// TIA Portal project "OPA_Demo" (V13)

(* hardware
DEVICE "S7-1200 station_1"  S7-1200 Station
   slot 0: "Rack_0"  Rack  V1.0
   slot 1: "PLC_1"  CPU 1214C DC/DC/DC  6ES7 214-1AG31-0XB0  V3.0
DEVICE "HMI_1"  KTP600 Basic color PN
   slot 0: "HMI"  HMI  6AV6 647-0AD11-3AX0  12.0.0.0
   slot 1: "HMI_RT_1"  KTP600 Basic color PN  6AV6 647-0AD11-3AX0  12.0.0.0
   slot 5: "HMI_1.IE_CP_1"  PROFINET Interface
      slot 1: "PROFINET Interface_1"  PROFINET Interface
         slot 1: "Port_1"  Port
*)

// ===== PLC "PLC_1"  CPU 1214C DC/DC/DC =====

VAR_GLOBAL   // PLC tag table "Input"
   "Tray_sensor" AT %I0.0 : Bool;
   "Doos_sensor" AT %I0.6 : Bool;
   "Tafel_sensor" AT %I0.4 : Bool;
   "Noodstop_aan_Plc" AT %I0.5 : Bool;
   "Noodstop_extern" AT %I0.3 : Bool;
   "Skip_Camera_Knop" AT %I0.1 : Bool;
   "Pause_Knop" AT %I0.2 : Bool;
END_VAR

VAR_GLOBAL   // PLC tag table "Memory"
   "HMI_Start_Pressed" AT %M42.0 : Bool;
   "HMI_Stop_Pressed" AT %M42.1 : Bool;
   "Running" AT %M42.2 : Bool;
   "HMI_White_Selected" AT %M42.3 : Bool;
   "HMI_Black_Pressed" AT %M42.4 : Bool;
   "HMI_tafel_omhoog" AT %M43.0 : Bool;
   "HMI_tafel_omlaag" AT %M43.1 : Bool;
   "HMI_tafel_inklappen" AT %M43.3 : Bool;
   "HMI_tafel_uitklappen" AT %M43.2 : Bool;
   "HMI_pneumatiek_aan" AT %M43.4 : Bool;
   "Noodstop" AT %M43.5 : Bool;
   "Noodrestart" AT %M43.6 : Bool;
   "Robot_TEMPORARY_BIT" AT %M43.7 : Bool;
   "Tafel_hoog" AT %M44.0 : Bool;
   "Noodstop_int" AT %MW50 : Int;
   "Next_Box_Ready" AT %M44.2 : Bool;
   "HardReset" AT %M44.3 : Bool;
   "Manual Mode" AT %M44.4 : Bool;
   "Pulse" AT %M44.5 : Bool;
   "Robot_Accepted" AT %M44.6 : Bool;
   "Camera_Box_Not_Empty" AT %M44.7 : Bool;
   "Placing_FIrst" AT %M45.0 : Bool;
   "Placing_Second" AT %M45.1 : Bool;
   "Camera_Not_Placed_Correctly" AT %M45.2 : Bool;
   "Waiting_For_Next_Order" AT %M45.3 : Bool;
   "Finished_Placing" AT %M45.4 : Bool;
   "Very Manual" AT %M45.5 : Bool;
   "Geen Robot Signaal" AT %M45.6 : Bool;
   "Tray_Found" AT %M45.7 : Bool;
   "Skip Camera" AT %M46.0 : Bool;
   "Paused" AT %M46.1 : Bool;
   "Start Running" AT %M46.2 : Bool;
END_VAR

VAR_GLOBAL   // PLC tag table "Output"
   "Tafel_uitklappen_cylinder" AT %Q0.1 : Bool;
   "Tafel_omhoog_cylinder" AT %Q0.4 : Bool;
   "Pneumatiek_aan" AT %Q0.2 : Bool;
   "Doosklem_Voor" AT %Q0.7 : Bool;
   "Doosklem_Achter" AT %Q0.5 : Bool;
   "VAN_ONDEREEEEEN!!!" AT %Q0.6 : Bool;
END_VAR

VAR_GLOBAL   // PLC tag table "Program Steps"
   "Waiting for Box" AT %M30.0 : Bool;
   "Box Arrived" AT %M30.1 : Bool;
   "Box Clamped" AT %M30.2 : Bool;
   "Preparing Table" AT %M31.0 : Bool;
   "Waiting for Robot" AT %M30.4 : Bool;
   "Robot is Finished" AT %M30.5 : Bool;
   "!LET HER RIP!" AT %M30.7 : Bool;
END_VAR

DATA_BLOCK "RobotConnectionDB"   // DB2
{ S7_Optimized_Access := 'FALSE' }
VERSION : 0.1
   VAR
      RobotAddress : TCON_IP_v4;
      Disconnect : Bool;
      ConnectID : Array[0..10] of UInt;
      BitWords : Array[0..1] of Word;
      Emergency_Stop : UInt;
      Run_Signal : UInt;
      Next_Box_ready : UInt;
      Stop_Register : UInt;
      Placing_Register : UInt;
      Finished_Placing_Register : UInt;
      Skip_Camera_Register : UInt;
      Done : Bool;
      Busy : Bool;
      Error : Bool;
      Status : Word;
      Statusses : Array[0..10] of Word;
      Stop_value : Word;
      Placing_value : Word;
      Finished_value : Word;
      Update_values : Bool;
   END_VAR
BEGIN
END_DATA_BLOCK

// folder: System blocks/Program resources

DATA_BLOCK "IEC_Timer_0_DB"   // DB1
{ S7_Optimized_Access := 'FALSE' }
AUTHOR : Simatic
FAMILY : IEC
NAME : IEC_TMR
VERSION : 1.0
// stored: InstanceOfName ?
"?"
BEGIN
END_DATA_BLOCK

DATA_BLOCK "IEC_Timer_0_DB_3"   // DB3
{ S7_Optimized_Access := 'FALSE' }
AUTHOR : Simatic
FAMILY : IEC
NAME : IEC_TMR
VERSION : 1.0
// stored: InstanceOfName ?
"?"
BEGIN
END_DATA_BLOCK

DATA_BLOCK "IEC_Timer_0_DB_4"   // DB7
{ S7_Optimized_Access := 'FALSE' }
AUTHOR : Simatic
FAMILY : IEC
NAME : IEC_TMR
VERSION : 1.0
// stored: InstanceOfName ?
"?"
BEGIN
END_DATA_BLOCK

DATA_BLOCK "IEC_Timer_0_DB_2"   // DB9
{ S7_Optimized_Access := 'FALSE' }
AUTHOR : Simatic
FAMILY : IEC
NAME : IEC_TMR
VERSION : 1.0
// stored: InstanceOfName ?
"?"
BEGIN
END_DATA_BLOCK

DATA_BLOCK "IEC_Timer_0_DB_6"   // DB14
{ S7_Optimized_Access := 'FALSE' }
AUTHOR : Simatic
FAMILY : IEC
NAME : IEC_TMR
VERSION : 1.0
// stored: InstanceOfName ?
"?"
BEGIN
END_DATA_BLOCK

DATA_BLOCK "IEC_Timer_0_DB_7"   // DB15
{ S7_Optimized_Access := 'FALSE' }
AUTHOR : Simatic
FAMILY : IEC
NAME : IEC_TMR
VERSION : 1.0
// stored: InstanceOfName ?
"?"
BEGIN
END_DATA_BLOCK

DATA_BLOCK "IEC_Timer_0_DB_8"   // DB16
{ S7_Optimized_Access := 'FALSE' }
AUTHOR : Simatic
FAMILY : IEC
NAME : IEC_TMR
VERSION : 1.0
// stored: InstanceOfName ?
"?"
BEGIN
END_DATA_BLOCK

DATA_BLOCK "IEC_Timer_0_DB_5"   // DB17
{ S7_Optimized_Access := 'FALSE' }
AUTHOR : Simatic
FAMILY : IEC
NAME : IEC_TMR
VERSION : 1.0
// stored: InstanceOfName ?
"?"
BEGIN
END_DATA_BLOCK

DATA_BLOCK "IEC_Timer_0_DB_9"   // DB18
{ S7_Optimized_Access := 'FALSE' }
AUTHOR : Simatic
FAMILY : IEC
NAME : IEC_TMR
VERSION : 1.0
// stored: InstanceOfName ?
"?"
BEGIN
END_DATA_BLOCK

DATA_BLOCK "IEC_Timer_0_DB_1"   // DB20
{ S7_Optimized_Access := 'FALSE' }
AUTHOR : Simatic
FAMILY : IEC
NAME : IEC_TMR
VERSION : 1.0
// stored: InstanceOfName ?
"?"
BEGIN
END_DATA_BLOCK

// folder: (top level)

FUNCTION "Program" : Void   // FC1, FBD
{ S7_Optimized_Access := 'FALSE' }
VERSION : 0.1
   VAR_TEMP   // added for the SCL form of the ladder/FBD networks
      _w1 : Bool;
      _w2 : Bool;
   END_VAR
BEGIN

REGION Network 1
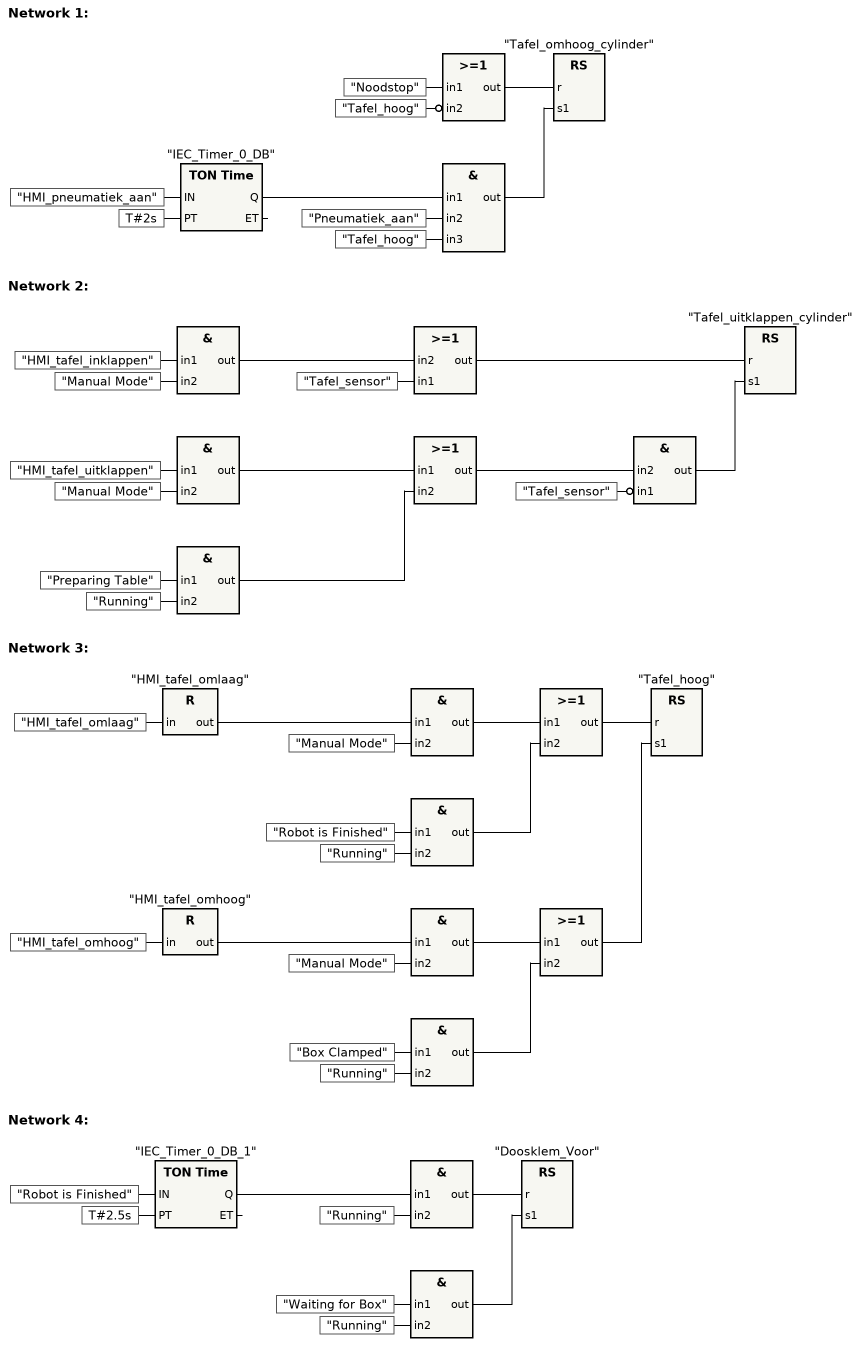
   "IEC_Timer_0_DB".TON(IN := "HMI_pneumatiek_aan", PT := T#2s);
   IF "Noodstop" OR NOT "Tafel_hoog" THEN
       "Tafel_omhoog_cylinder" := FALSE;   // RS flip-flop
   END_IF;
   IF "IEC_Timer_0_DB".Q AND "Pneumatiek_aan" AND "Tafel_hoog" THEN "Tafel_omhoog_cylinder" := TRUE; END_IF;
END_REGION

REGION Network 2
   IF ("HMI_tafel_inklappen" AND "Manual Mode") OR "Tafel_sensor" THEN
       "Tafel_uitklappen_cylinder" := FALSE;   // RS flip-flop
   END_IF;
   IF (("HMI_tafel_uitklappen" AND "Manual Mode") OR ("Preparing Table" AND "Running")) AND NOT "Tafel_sensor" THEN
       "Tafel_uitklappen_cylinder" := TRUE;
   END_IF;
END_REGION

REGION Network 3
   #_w1 := "HMI_tafel_omlaag";
   IF #_w1 THEN "HMI_tafel_omlaag" := FALSE; END_IF;
   #_w2 := "HMI_tafel_omhoog";
   IF #_w2 THEN "HMI_tafel_omhoog" := FALSE; END_IF;
   IF (#_w1 AND "Manual Mode") OR ("Robot is Finished" AND "Running") THEN
       "Tafel_hoog" := FALSE;   // RS flip-flop
   END_IF;
   IF (#_w2 AND "Manual Mode") OR ("Box Clamped" AND "Running") THEN "Tafel_hoog" := TRUE; END_IF;
END_REGION

REGION Network 4
   "IEC_Timer_0_DB_1".TON(IN := "Robot is Finished", PT := T#2.5s);
   IF "IEC_Timer_0_DB_1".Q AND "Running" THEN
       "Doosklem_Voor" := FALSE;   // RS flip-flop
   END_IF;
   IF "Waiting for Box" AND "Running" THEN "Doosklem_Voor" := TRUE; END_IF;
END_REGION

REGION Network 5
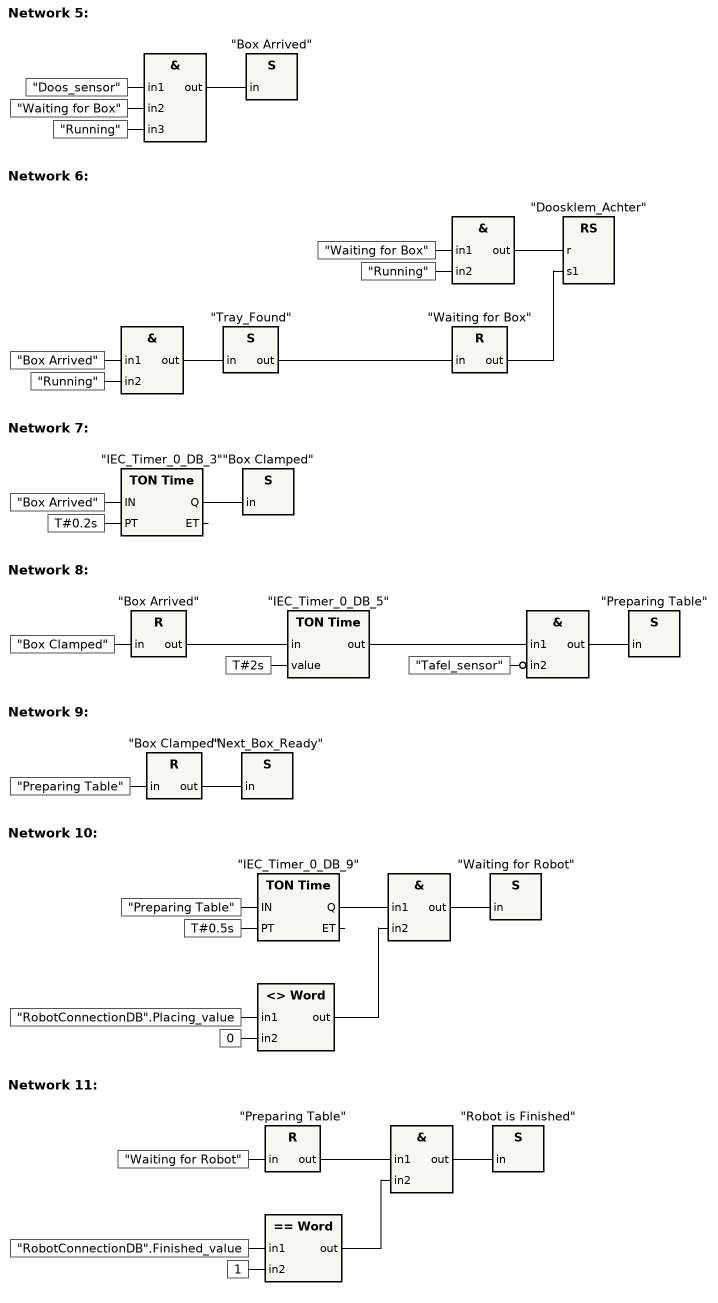
   IF "Doos_sensor" AND "Waiting for Box" AND "Running" THEN "Box Arrived" := TRUE; END_IF;
END_REGION

REGION Network 6
   #_w1 := "Box Arrived" AND "Running";
   IF #_w1 THEN "Tray_Found" := TRUE; END_IF;
   #_w2 := "Waiting for Box" AND "Running";
   IF #_w1 THEN "Waiting for Box" := FALSE; END_IF;
   IF #_w2 THEN
       "Doosklem_Achter" := FALSE;   // RS flip-flop
   END_IF;
   IF #_w1 THEN "Doosklem_Achter" := TRUE; END_IF;
END_REGION

REGION Network 7
   "IEC_Timer_0_DB_3".TON(IN := "Box Arrived", PT := T#0.2s);
   IF "IEC_Timer_0_DB_3".Q THEN "Box Clamped" := TRUE; END_IF;
END_REGION

REGION Network 8
   IF "Box Clamped" THEN "Box Arrived" := FALSE; END_IF;
   "IEC_Timer_0_DB_5".TON(IN := "Box Clamped", PT := T#2s);   // TON coil
   IF "Box Clamped" AND NOT "Tafel_sensor" THEN "Preparing Table" := TRUE; END_IF;
END_REGION

REGION Network 9
   IF "Preparing Table" THEN
       "Box Clamped" := FALSE;
       "Next_Box_Ready" := TRUE;
   END_IF;
END_REGION

REGION Network 10
   "IEC_Timer_0_DB_9".TON(IN := "Preparing Table", PT := T#0.5s);
   IF "IEC_Timer_0_DB_9".Q AND ("RobotConnectionDB".Placing_value <> 0) THEN
       "Waiting for Robot" := TRUE;
   END_IF;
END_REGION

REGION Network 11
   IF "Waiting for Robot" THEN "Preparing Table" := FALSE; END_IF;
   IF "Waiting for Robot" AND ("RobotConnectionDB".Finished_value = 1) THEN
       "Robot is Finished" := TRUE;
   END_IF;
END_REGION

REGION Network 12
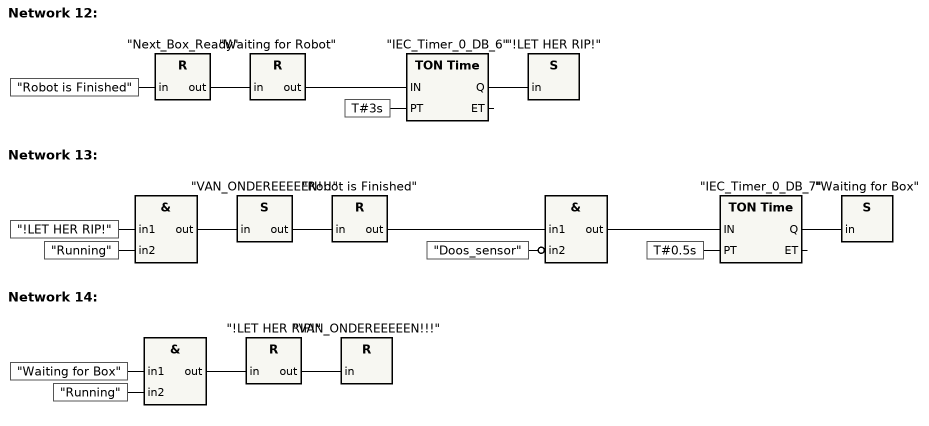
   IF "Robot is Finished" THEN
       "Next_Box_Ready" := FALSE;
       "Waiting for Robot" := FALSE;
   END_IF;
   "IEC_Timer_0_DB_6".TON(IN := "Robot is Finished", PT := T#3s);
   IF "IEC_Timer_0_DB_6".Q THEN "!LET HER RIP!" := TRUE; END_IF;
END_REGION

REGION Network 13
   #_w1 := "!LET HER RIP!" AND "Running";
   IF #_w1 THEN
       "VAN_ONDEREEEEEN!!!" := TRUE;
       "Robot is Finished" := FALSE;
   END_IF;
   "IEC_Timer_0_DB_7".TON(IN := #_w1 AND NOT "Doos_sensor", PT := T#0.5s);
   IF "IEC_Timer_0_DB_7".Q THEN "Waiting for Box" := TRUE; END_IF;
END_REGION

REGION Network 14
   IF "Waiting for Box" AND "Running" THEN
       "!LET HER RIP!" := FALSE;
       "VAN_ONDEREEEEEN!!!" := FALSE;
   END_IF;
END_REGION
END_FUNCTION

FUNCTION "Set_Noodstop" : Void   // FC2, SCL
{ S7_Optimized_Access := 'FALSE' }
VERSION : 0.1
BEGIN
   IF "Noodstop" THEN
       // Statement section IF
       "Noodstop_int" := 4;
       ;
   ELSE
       "Noodstop_int" := 0;
       ;
   END_IF;
END_FUNCTION

FUNCTION "RobotConnection" : Void   // FC3, FBD
{ S7_Optimized_Access := 'FALSE' }
VERSION : 0.1
BEGIN

REGION Network 1
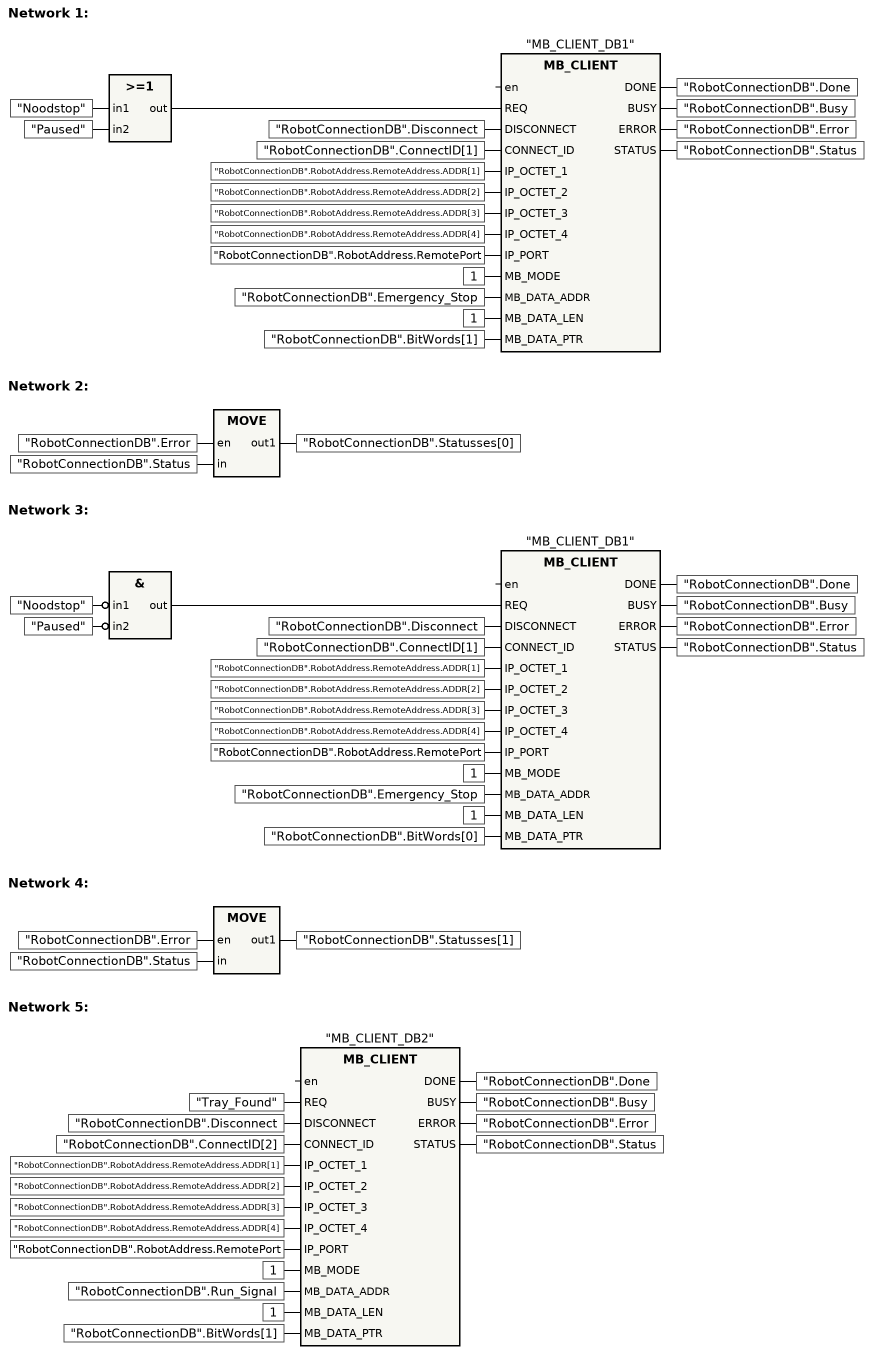
   "MB_CLIENT_DB1"(REQ := "Noodstop" OR "Paused",   // MB_CLIENT
                   DISCONNECT := "RobotConnectionDB".Disconnect,
                   CONNECT_ID := "RobotConnectionDB".ConnectID[1],
                   IP_OCTET_1 := "RobotConnectionDB".RobotAddress.RemoteAddress.ADDR[1],
                   IP_OCTET_2 := "RobotConnectionDB".RobotAddress.RemoteAddress.ADDR[2],
                   IP_OCTET_3 := "RobotConnectionDB".RobotAddress.RemoteAddress.ADDR[3],
                   IP_OCTET_4 := "RobotConnectionDB".RobotAddress.RemoteAddress.ADDR[4],
                   IP_PORT := "RobotConnectionDB".RobotAddress.RemotePort,
                   MB_MODE := 1,
                   MB_DATA_ADDR := "RobotConnectionDB".Emergency_Stop,
                   MB_DATA_LEN := 1,
                   MB_DATA_PTR := "RobotConnectionDB".BitWords[1],
                   DONE => "RobotConnectionDB".Done,
                   BUSY => "RobotConnectionDB".Busy,
                   ERROR => "RobotConnectionDB".Error,
                   STATUS => "RobotConnectionDB".Status);
END_REGION

REGION Network 2
   IF "RobotConnectionDB".Error THEN "RobotConnectionDB".Statusses[0] := "RobotConnectionDB".Status; END_IF;
END_REGION

REGION Network 3
   "MB_CLIENT_DB1"(REQ := NOT "Noodstop" AND NOT "Paused",   // MB_CLIENT
                   DISCONNECT := "RobotConnectionDB".Disconnect,
                   CONNECT_ID := "RobotConnectionDB".ConnectID[1],
                   IP_OCTET_1 := "RobotConnectionDB".RobotAddress.RemoteAddress.ADDR[1],
                   IP_OCTET_2 := "RobotConnectionDB".RobotAddress.RemoteAddress.ADDR[2],
                   IP_OCTET_3 := "RobotConnectionDB".RobotAddress.RemoteAddress.ADDR[3],
                   IP_OCTET_4 := "RobotConnectionDB".RobotAddress.RemoteAddress.ADDR[4],
                   IP_PORT := "RobotConnectionDB".RobotAddress.RemotePort,
                   MB_MODE := 1,
                   MB_DATA_ADDR := "RobotConnectionDB".Emergency_Stop,
                   MB_DATA_LEN := 1,
                   MB_DATA_PTR := "RobotConnectionDB".BitWords[0],
                   DONE => "RobotConnectionDB".Done,
                   BUSY => "RobotConnectionDB".Busy,
                   ERROR => "RobotConnectionDB".Error,
                   STATUS => "RobotConnectionDB".Status);
END_REGION

REGION Network 4
   IF "RobotConnectionDB".Error THEN "RobotConnectionDB".Statusses[1] := "RobotConnectionDB".Status; END_IF;
END_REGION

REGION Network 5
   "MB_CLIENT_DB2"(REQ := "Tray_Found",   // MB_CLIENT
                   DISCONNECT := "RobotConnectionDB".Disconnect,
                   CONNECT_ID := "RobotConnectionDB".ConnectID[2],
                   IP_OCTET_1 := "RobotConnectionDB".RobotAddress.RemoteAddress.ADDR[1],
                   IP_OCTET_2 := "RobotConnectionDB".RobotAddress.RemoteAddress.ADDR[2],
                   IP_OCTET_3 := "RobotConnectionDB".RobotAddress.RemoteAddress.ADDR[3],
                   IP_OCTET_4 := "RobotConnectionDB".RobotAddress.RemoteAddress.ADDR[4],
                   IP_PORT := "RobotConnectionDB".RobotAddress.RemotePort,
                   MB_MODE := 1,
                   MB_DATA_ADDR := "RobotConnectionDB".Run_Signal,
                   MB_DATA_LEN := 1,
                   MB_DATA_PTR := "RobotConnectionDB".BitWords[1],
                   DONE => "RobotConnectionDB".Done,
                   BUSY => "RobotConnectionDB".Busy,
                   ERROR => "RobotConnectionDB".Error,
                   STATUS => "RobotConnectionDB".Status);
END_REGION

REGION Network 6
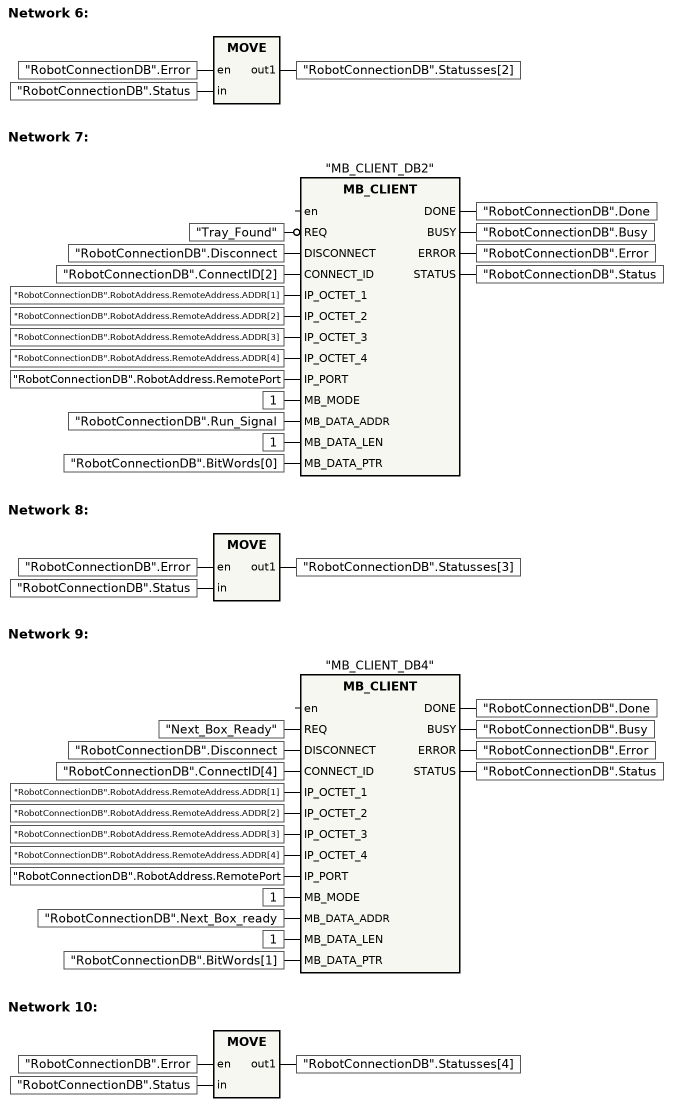
   IF "RobotConnectionDB".Error THEN "RobotConnectionDB".Statusses[2] := "RobotConnectionDB".Status; END_IF;
END_REGION

REGION Network 7
   "MB_CLIENT_DB2"(REQ := NOT "Tray_Found",   // MB_CLIENT
                   DISCONNECT := "RobotConnectionDB".Disconnect,
                   CONNECT_ID := "RobotConnectionDB".ConnectID[2],
                   IP_OCTET_1 := "RobotConnectionDB".RobotAddress.RemoteAddress.ADDR[1],
                   IP_OCTET_2 := "RobotConnectionDB".RobotAddress.RemoteAddress.ADDR[2],
                   IP_OCTET_3 := "RobotConnectionDB".RobotAddress.RemoteAddress.ADDR[3],
                   IP_OCTET_4 := "RobotConnectionDB".RobotAddress.RemoteAddress.ADDR[4],
                   IP_PORT := "RobotConnectionDB".RobotAddress.RemotePort,
                   MB_MODE := 1,
                   MB_DATA_ADDR := "RobotConnectionDB".Run_Signal,
                   MB_DATA_LEN := 1,
                   MB_DATA_PTR := "RobotConnectionDB".BitWords[0],
                   DONE => "RobotConnectionDB".Done,
                   BUSY => "RobotConnectionDB".Busy,
                   ERROR => "RobotConnectionDB".Error,
                   STATUS => "RobotConnectionDB".Status);
END_REGION

REGION Network 8
   IF "RobotConnectionDB".Error THEN "RobotConnectionDB".Statusses[3] := "RobotConnectionDB".Status; END_IF;
END_REGION

REGION Network 9
   "MB_CLIENT_DB4"(REQ := "Next_Box_Ready",   // MB_CLIENT
                   DISCONNECT := "RobotConnectionDB".Disconnect,
                   CONNECT_ID := "RobotConnectionDB".ConnectID[4],
                   IP_OCTET_1 := "RobotConnectionDB".RobotAddress.RemoteAddress.ADDR[1],
                   IP_OCTET_2 := "RobotConnectionDB".RobotAddress.RemoteAddress.ADDR[2],
                   IP_OCTET_3 := "RobotConnectionDB".RobotAddress.RemoteAddress.ADDR[3],
                   IP_OCTET_4 := "RobotConnectionDB".RobotAddress.RemoteAddress.ADDR[4],
                   IP_PORT := "RobotConnectionDB".RobotAddress.RemotePort,
                   MB_MODE := 1,
                   MB_DATA_ADDR := "RobotConnectionDB".Next_Box_ready,
                   MB_DATA_LEN := 1,
                   MB_DATA_PTR := "RobotConnectionDB".BitWords[1],
                   DONE => "RobotConnectionDB".Done,
                   BUSY => "RobotConnectionDB".Busy,
                   ERROR => "RobotConnectionDB".Error,
                   STATUS => "RobotConnectionDB".Status);
END_REGION

REGION Network 10
   IF "RobotConnectionDB".Error THEN "RobotConnectionDB".Statusses[4] := "RobotConnectionDB".Status; END_IF;
END_REGION

REGION Network 11
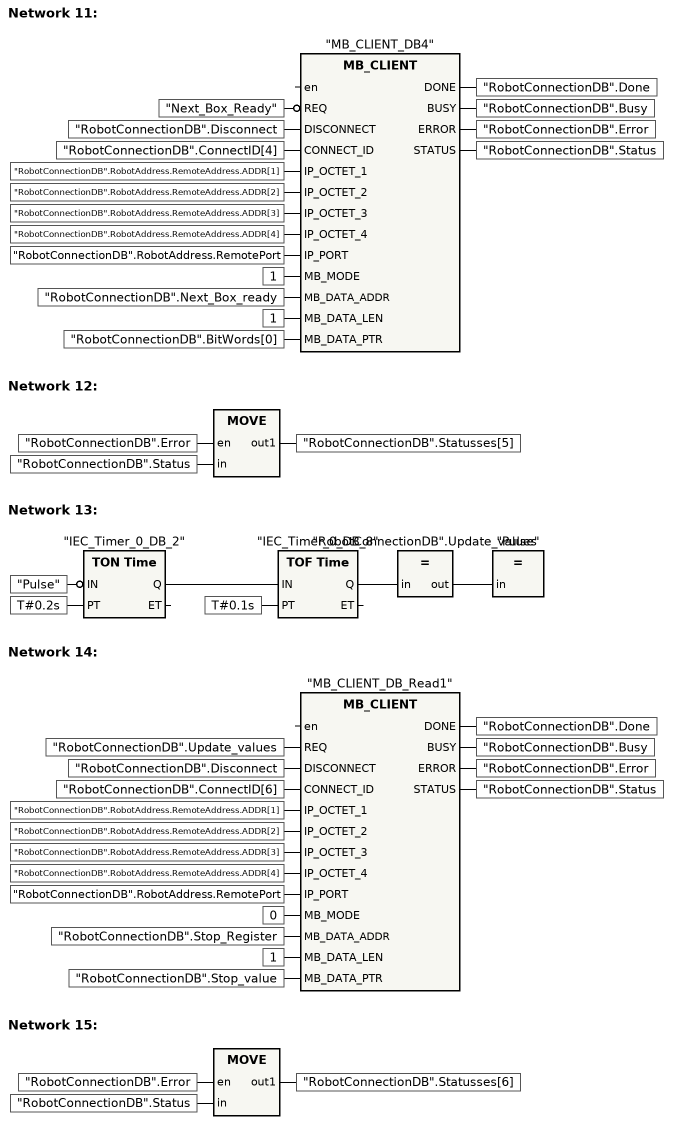
   "MB_CLIENT_DB4"(REQ := NOT "Next_Box_Ready",   // MB_CLIENT
                   DISCONNECT := "RobotConnectionDB".Disconnect,
                   CONNECT_ID := "RobotConnectionDB".ConnectID[4],
                   IP_OCTET_1 := "RobotConnectionDB".RobotAddress.RemoteAddress.ADDR[1],
                   IP_OCTET_2 := "RobotConnectionDB".RobotAddress.RemoteAddress.ADDR[2],
                   IP_OCTET_3 := "RobotConnectionDB".RobotAddress.RemoteAddress.ADDR[3],
                   IP_OCTET_4 := "RobotConnectionDB".RobotAddress.RemoteAddress.ADDR[4],
                   IP_PORT := "RobotConnectionDB".RobotAddress.RemotePort,
                   MB_MODE := 1,
                   MB_DATA_ADDR := "RobotConnectionDB".Next_Box_ready,
                   MB_DATA_LEN := 1,
                   MB_DATA_PTR := "RobotConnectionDB".BitWords[0],
                   DONE => "RobotConnectionDB".Done,
                   BUSY => "RobotConnectionDB".Busy,
                   ERROR => "RobotConnectionDB".Error,
                   STATUS => "RobotConnectionDB".Status);
END_REGION

REGION Network 12
   IF "RobotConnectionDB".Error THEN "RobotConnectionDB".Statusses[5] := "RobotConnectionDB".Status; END_IF;
END_REGION

REGION Network 13
   "IEC_Timer_0_DB_2".TON(IN := NOT "Pulse", PT := T#0.2s);
   "IEC_Timer_0_DB_8".TOF(IN := "IEC_Timer_0_DB_2".Q, PT := T#0.1s);
   "RobotConnectionDB".Update_values := "IEC_Timer_0_DB_8".Q;
   "Pulse" := "IEC_Timer_0_DB_8".Q;
END_REGION

REGION Network 14
   "MB_CLIENT_DB_Read1"(REQ := "RobotConnectionDB".Update_values,   // MB_CLIENT
                        DISCONNECT := "RobotConnectionDB".Disconnect,
                        CONNECT_ID := "RobotConnectionDB".ConnectID[6],
                        IP_OCTET_1 := "RobotConnectionDB".RobotAddress.RemoteAddress.ADDR[1],
                        IP_OCTET_2 := "RobotConnectionDB".RobotAddress.RemoteAddress.ADDR[2],
                        IP_OCTET_3 := "RobotConnectionDB".RobotAddress.RemoteAddress.ADDR[3],
                        IP_OCTET_4 := "RobotConnectionDB".RobotAddress.RemoteAddress.ADDR[4],
                        IP_PORT := "RobotConnectionDB".RobotAddress.RemotePort,
                        MB_MODE := 0,
                        MB_DATA_ADDR := "RobotConnectionDB".Stop_Register,
                        MB_DATA_LEN := 1,
                        MB_DATA_PTR := "RobotConnectionDB".Stop_value,
                        DONE => "RobotConnectionDB".Done,
                        BUSY => "RobotConnectionDB".Busy,
                        ERROR => "RobotConnectionDB".Error,
                        STATUS => "RobotConnectionDB".Status);
END_REGION

REGION Network 15
   IF "RobotConnectionDB".Error THEN "RobotConnectionDB".Statusses[6] := "RobotConnectionDB".Status; END_IF;
END_REGION

REGION Network 16
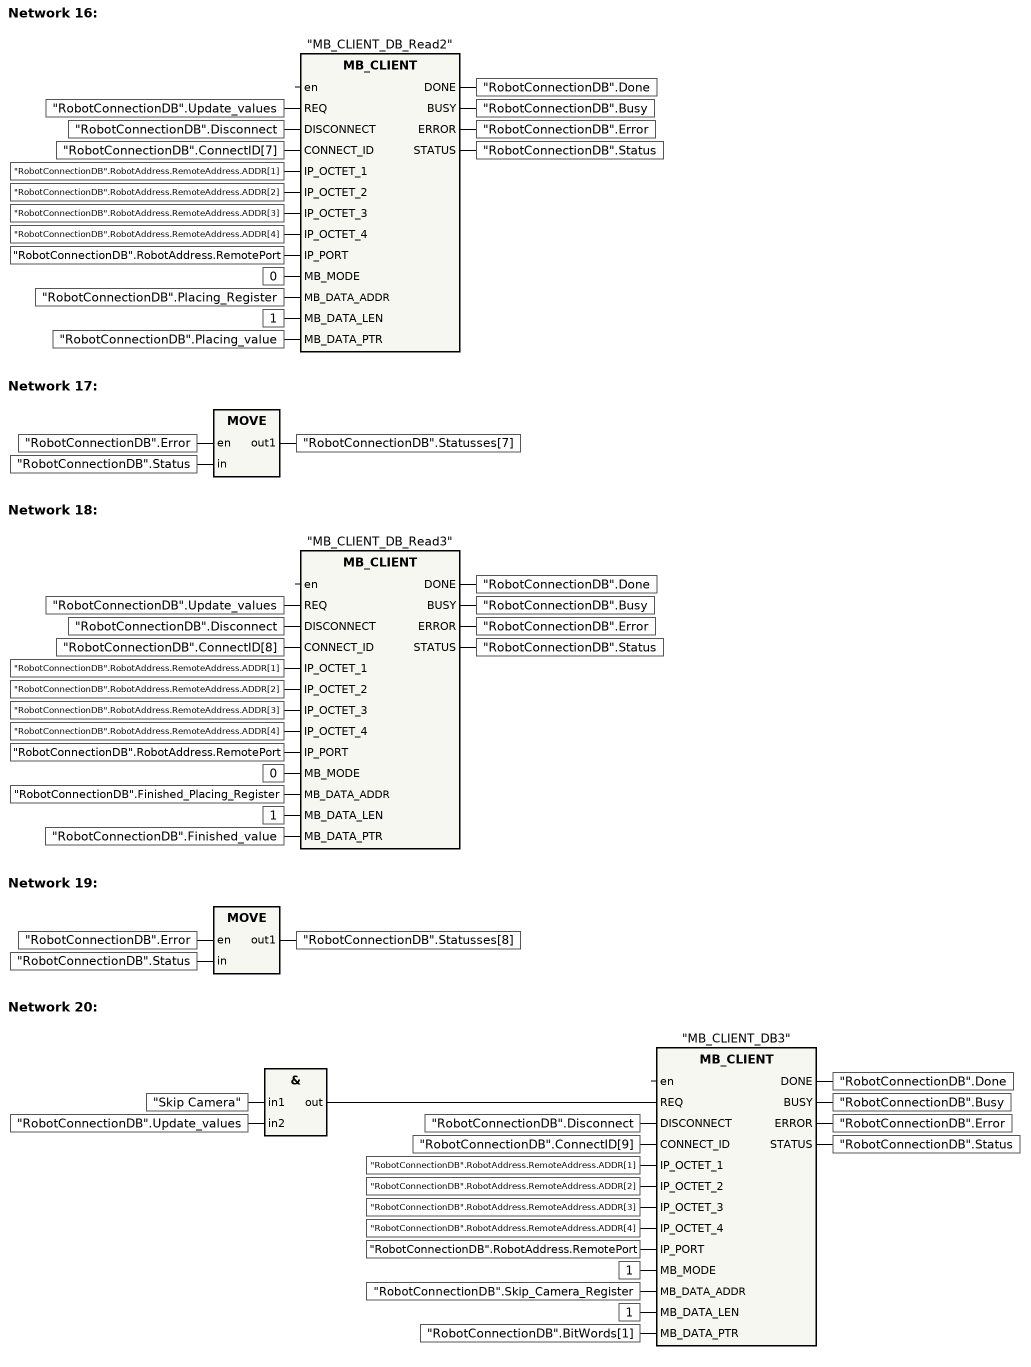
   "MB_CLIENT_DB_Read2"(REQ := "RobotConnectionDB".Update_values,   // MB_CLIENT
                        DISCONNECT := "RobotConnectionDB".Disconnect,
                        CONNECT_ID := "RobotConnectionDB".ConnectID[7],
                        IP_OCTET_1 := "RobotConnectionDB".RobotAddress.RemoteAddress.ADDR[1],
                        IP_OCTET_2 := "RobotConnectionDB".RobotAddress.RemoteAddress.ADDR[2],
                        IP_OCTET_3 := "RobotConnectionDB".RobotAddress.RemoteAddress.ADDR[3],
                        IP_OCTET_4 := "RobotConnectionDB".RobotAddress.RemoteAddress.ADDR[4],
                        IP_PORT := "RobotConnectionDB".RobotAddress.RemotePort,
                        MB_MODE := 0,
                        MB_DATA_ADDR := "RobotConnectionDB".Placing_Register,
                        MB_DATA_LEN := 1,
                        MB_DATA_PTR := "RobotConnectionDB".Placing_value,
                        DONE => "RobotConnectionDB".Done,
                        BUSY => "RobotConnectionDB".Busy,
                        ERROR => "RobotConnectionDB".Error,
                        STATUS => "RobotConnectionDB".Status);
END_REGION

REGION Network 17
   IF "RobotConnectionDB".Error THEN "RobotConnectionDB".Statusses[7] := "RobotConnectionDB".Status; END_IF;
END_REGION

REGION Network 18
   "MB_CLIENT_DB_Read3"(REQ := "RobotConnectionDB".Update_values,   // MB_CLIENT
                        DISCONNECT := "RobotConnectionDB".Disconnect,
                        CONNECT_ID := "RobotConnectionDB".ConnectID[8],
                        IP_OCTET_1 := "RobotConnectionDB".RobotAddress.RemoteAddress.ADDR[1],
                        IP_OCTET_2 := "RobotConnectionDB".RobotAddress.RemoteAddress.ADDR[2],
                        IP_OCTET_3 := "RobotConnectionDB".RobotAddress.RemoteAddress.ADDR[3],
                        IP_OCTET_4 := "RobotConnectionDB".RobotAddress.RemoteAddress.ADDR[4],
                        IP_PORT := "RobotConnectionDB".RobotAddress.RemotePort,
                        MB_MODE := 0,
                        MB_DATA_ADDR := "RobotConnectionDB".Finished_Placing_Register,
                        MB_DATA_LEN := 1,
                        MB_DATA_PTR := "RobotConnectionDB".Finished_value,
                        DONE => "RobotConnectionDB".Done,
                        BUSY => "RobotConnectionDB".Busy,
                        ERROR => "RobotConnectionDB".Error,
                        STATUS => "RobotConnectionDB".Status);
END_REGION

REGION Network 19
   IF "RobotConnectionDB".Error THEN "RobotConnectionDB".Statusses[8] := "RobotConnectionDB".Status; END_IF;
END_REGION

REGION Network 20
   "MB_CLIENT_DB3"(REQ := "Skip Camera" AND "RobotConnectionDB".Update_values,   // MB_CLIENT
                   DISCONNECT := "RobotConnectionDB".Disconnect,
                   CONNECT_ID := "RobotConnectionDB".ConnectID[9],
                   IP_OCTET_1 := "RobotConnectionDB".RobotAddress.RemoteAddress.ADDR[1],
                   IP_OCTET_2 := "RobotConnectionDB".RobotAddress.RemoteAddress.ADDR[2],
                   IP_OCTET_3 := "RobotConnectionDB".RobotAddress.RemoteAddress.ADDR[3],
                   IP_OCTET_4 := "RobotConnectionDB".RobotAddress.RemoteAddress.ADDR[4],
                   IP_PORT := "RobotConnectionDB".RobotAddress.RemotePort,
                   MB_MODE := 1,
                   MB_DATA_ADDR := "RobotConnectionDB".Skip_Camera_Register,
                   MB_DATA_LEN := 1,
                   MB_DATA_PTR := "RobotConnectionDB".BitWords[1],
                   DONE => "RobotConnectionDB".Done,
                   BUSY => "RobotConnectionDB".Busy,
                   ERROR => "RobotConnectionDB".Error,
                   STATUS => "RobotConnectionDB".Status);
END_REGION

REGION Network 21
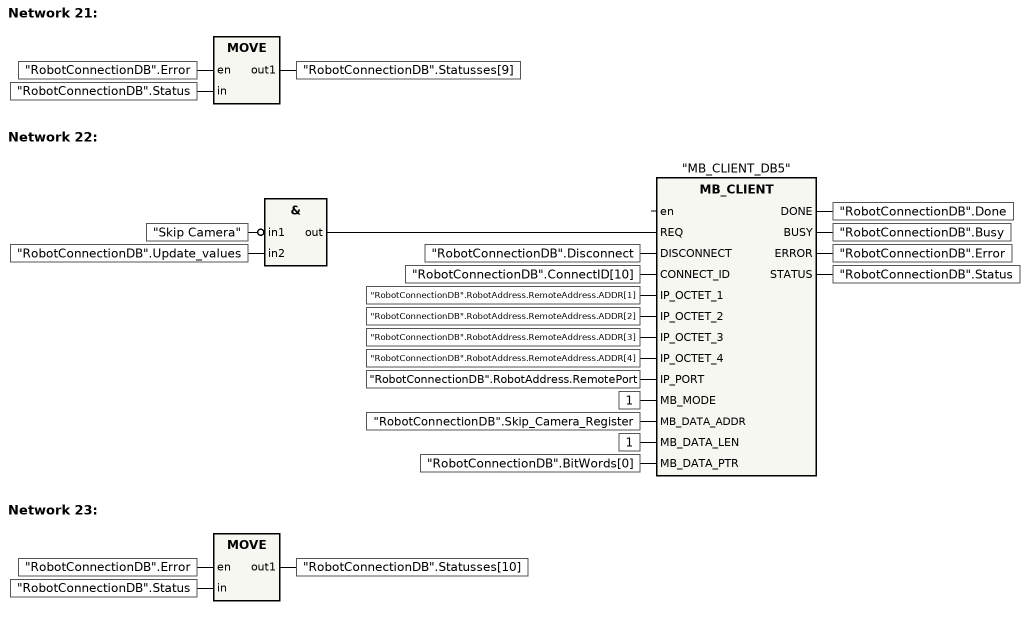
   IF "RobotConnectionDB".Error THEN "RobotConnectionDB".Statusses[9] := "RobotConnectionDB".Status; END_IF;
END_REGION

REGION Network 22
   "MB_CLIENT_DB5"(REQ := NOT "Skip Camera" AND "RobotConnectionDB".Update_values,   // MB_CLIENT
                   DISCONNECT := "RobotConnectionDB".Disconnect,
                   CONNECT_ID := "RobotConnectionDB".ConnectID[10],
                   IP_OCTET_1 := "RobotConnectionDB".RobotAddress.RemoteAddress.ADDR[1],
                   IP_OCTET_2 := "RobotConnectionDB".RobotAddress.RemoteAddress.ADDR[2],
                   IP_OCTET_3 := "RobotConnectionDB".RobotAddress.RemoteAddress.ADDR[3],
                   IP_OCTET_4 := "RobotConnectionDB".RobotAddress.RemoteAddress.ADDR[4],
                   IP_PORT := "RobotConnectionDB".RobotAddress.RemotePort,
                   MB_MODE := 1,
                   MB_DATA_ADDR := "RobotConnectionDB".Skip_Camera_Register,
                   MB_DATA_LEN := 1,
                   MB_DATA_PTR := "RobotConnectionDB".BitWords[0],
                   DONE => "RobotConnectionDB".Done,
                   BUSY => "RobotConnectionDB".Busy,
                   ERROR => "RobotConnectionDB".Error,
                   STATUS => "RobotConnectionDB".Status);
END_REGION

REGION Network 23
   IF "RobotConnectionDB".Error THEN "RobotConnectionDB".Statusses[10] := "RobotConnectionDB".Status; END_IF;
END_REGION
END_FUNCTION

FUNCTION "Reset" : Void   // FC4, SCL
{ S7_Optimized_Access := 'FALSE' }
VERSION : 0.1
BEGIN
   //Set Outputs to zero
   "Tafel_uitklappen_cylinder" := 0;
   "Tafel_omhoog_cylinder" := 0;
   "Pneumatiek_aan" := 0;
   "Doosklem_Voor" := 0;
   "Doosklem_Achter" := 0;
   "VAN_ONDEREEEEEN!!!" := 0;

   //Prepare Memory
   "Running" := 0;
   "Noodrestart" := 0;
   "Tafel_hoog" := 0;
   "Next_Box_Ready" := 0;
   "Tray_Found" := 0;
   "Skip Camera" := 0;

   //Prepare Program Steps
   "Waiting for Box" := 1;
   "Box Arrived" := 0;
   "Box Clamped" := 0;
   "Preparing Table" := 0;
   "Waiting for Robot" := 0;
   "Robot is Finished" := 0;
   "!LET HER RIP!" := 0;
END_FUNCTION

FUNCTION "Status_Update" : Void   // FC5, FBD
{ S7_Optimized_Access := 'FALSE' }
VERSION : 0.1
BEGIN

REGION Network 1
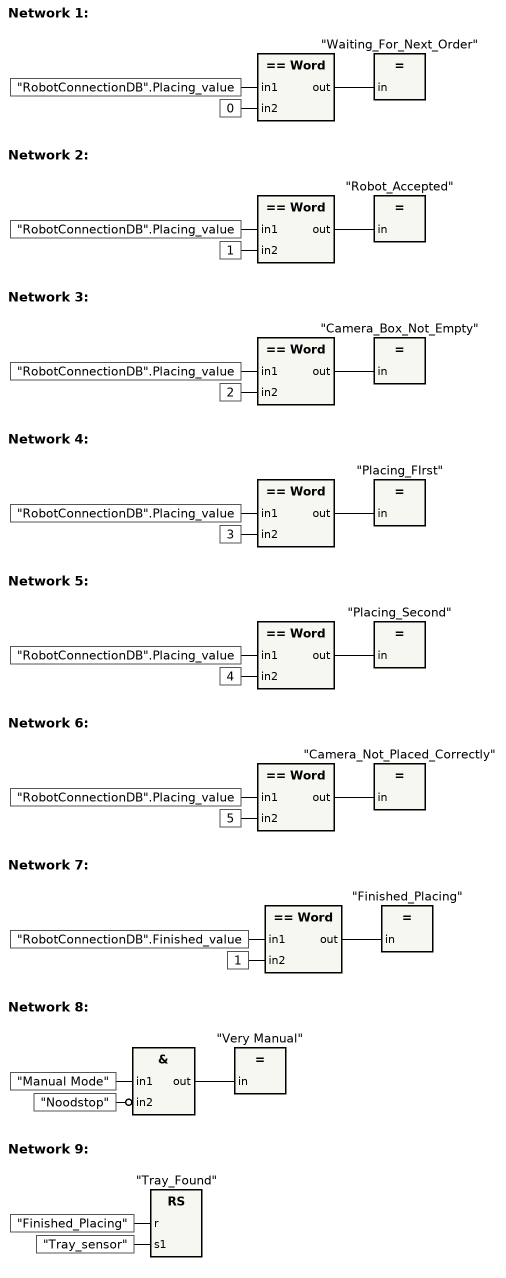
   "Waiting_For_Next_Order" := "RobotConnectionDB".Placing_value = 0;
END_REGION

REGION Network 2
   "Robot_Accepted" := "RobotConnectionDB".Placing_value = 1;
END_REGION

REGION Network 3
   "Camera_Box_Not_Empty" := "RobotConnectionDB".Placing_value = 2;
END_REGION

REGION Network 4
   "Placing_FIrst" := "RobotConnectionDB".Placing_value = 3;
END_REGION

REGION Network 5
   "Placing_Second" := "RobotConnectionDB".Placing_value = 4;
END_REGION

REGION Network 6
   "Camera_Not_Placed_Correctly" := "RobotConnectionDB".Placing_value = 5;
END_REGION

REGION Network 7
   "Finished_Placing" := "RobotConnectionDB".Finished_value = 1;
END_REGION

REGION Network 8
   "Very Manual" := "Manual Mode" AND NOT "Noodstop";
END_REGION

REGION Network 9
   IF "Finished_Placing" THEN
       "Tray_Found" := FALSE;   // RS flip-flop
   END_IF;
   IF "Tray_sensor" THEN "Tray_Found" := TRUE; END_IF;
END_REGION

REGION Network 10
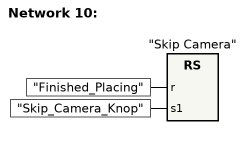
   IF "Finished_Placing" THEN
       "Skip Camera" := FALSE;   // RS flip-flop
   END_IF;
   IF "Skip_Camera_Knop" THEN "Skip Camera" := TRUE; END_IF;
END_REGION
END_FUNCTION

FUNCTION "Reset_Program_Steps" : Void   // FC6, SCL
{ S7_Optimized_Access := 'FALSE' }
VERSION : 0.1
BEGIN
   //Prepare Program Steps
   "Waiting for Box" := 1;
   "Box Arrived" := 0;
   "Box Clamped" := 0;
   "Preparing Table" := 0;
   "Waiting for Robot" := 0;
   "Robot is Finished" := 0;
   "!LET HER RIP!" := 0;
END_FUNCTION

ORGANIZATION_BLOCK "Main"   // OB1, FBD, ProgramCycle
TITLE = "Main Program Sweep (Cycle)"
{ S7_Optimized_Access := 'FALSE' }
VERSION : 0.1
   VAR_TEMP   // added for the SCL form of the ladder/FBD networks
      _w1 : Bool;
      _w2 : Bool;
      _w3 : Bool;
   END_VAR
BEGIN

REGION Network 1
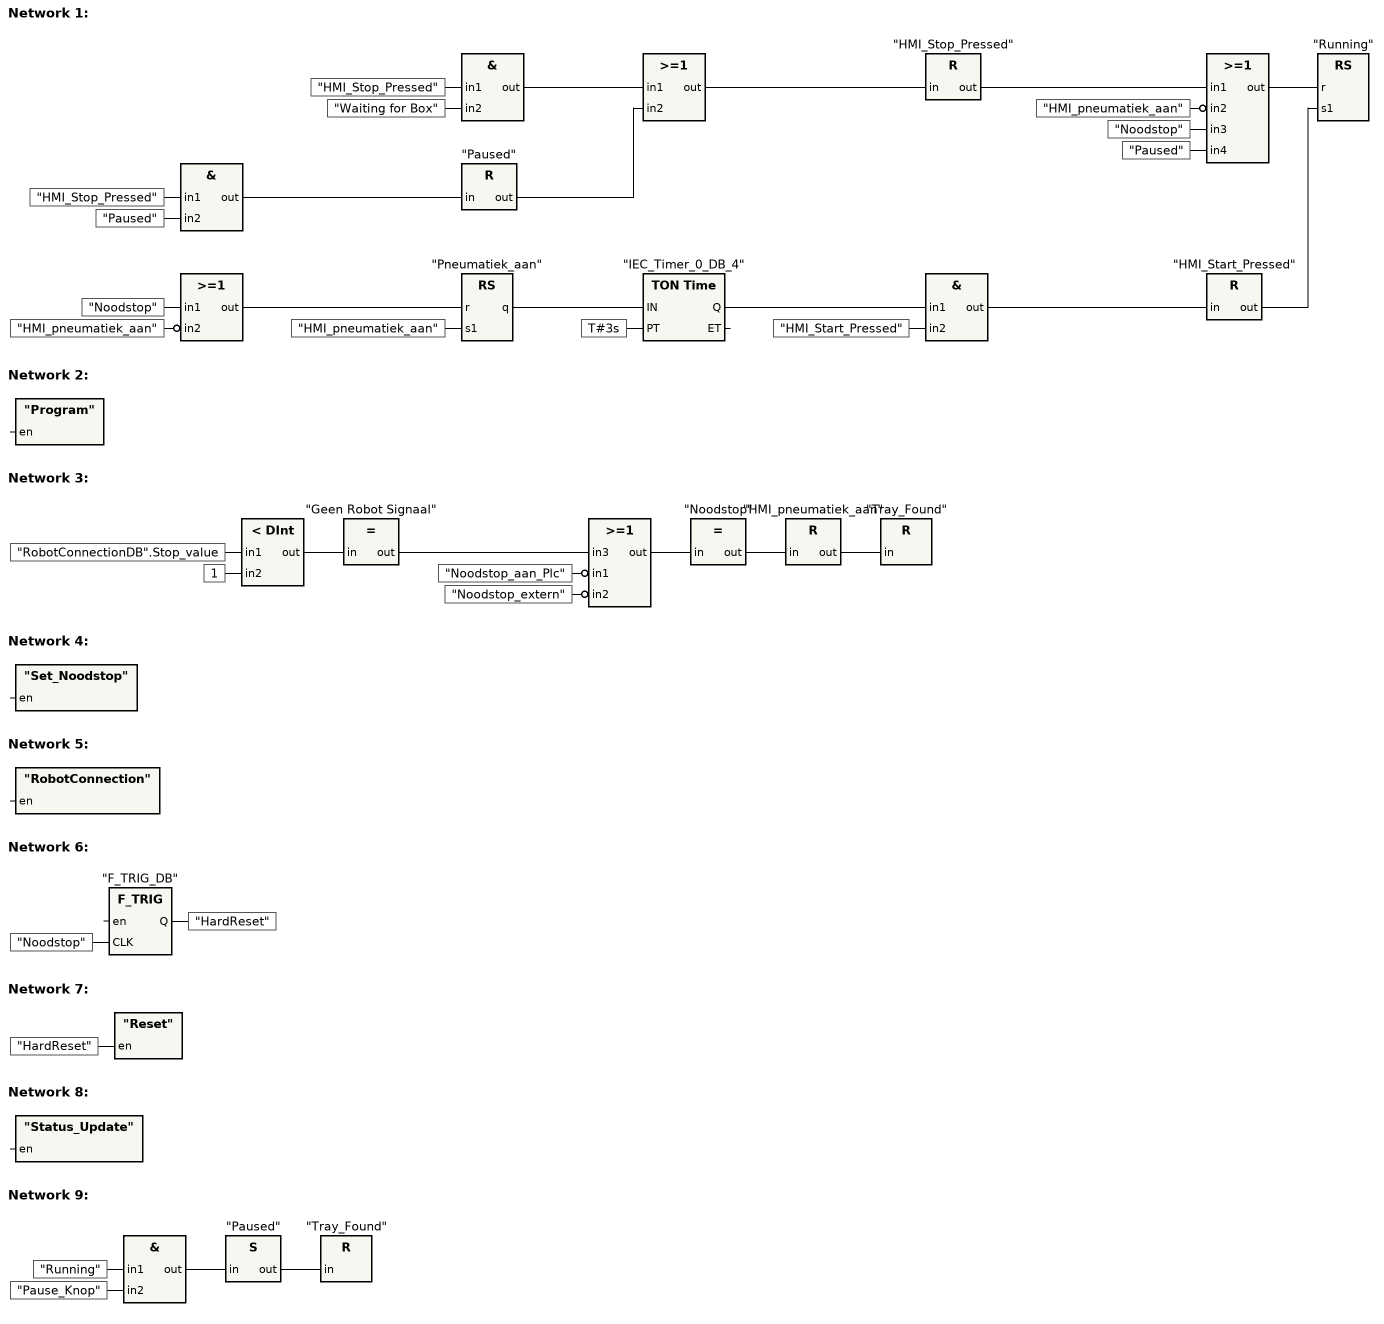
   #_w1 := "HMI_Stop_Pressed" AND "Paused";
   IF #_w1 THEN "Paused" := FALSE; END_IF;
   #_w2 := ("HMI_Stop_Pressed" AND "Waiting for Box") OR #_w1;
   IF #_w2 THEN "HMI_Stop_Pressed" := FALSE; END_IF;
   IF "Noodstop" OR NOT "HMI_pneumatiek_aan" THEN
       "Pneumatiek_aan" := FALSE;   // RS flip-flop
   END_IF;
   IF "HMI_pneumatiek_aan" THEN "Pneumatiek_aan" := TRUE; END_IF;
   "IEC_Timer_0_DB_4".TON(IN := "Pneumatiek_aan", PT := T#3s);
   #_w3 := "IEC_Timer_0_DB_4".Q AND "HMI_Start_Pressed";
   IF #_w3 THEN "HMI_Start_Pressed" := FALSE; END_IF;
   IF #_w2 OR NOT "HMI_pneumatiek_aan" OR "Noodstop" OR "Paused" THEN
       "Running" := FALSE;   // RS flip-flop
   END_IF;
   IF #_w3 THEN "Running" := TRUE; END_IF;
END_REGION

REGION Network 2
   "Program"();
END_REGION

REGION Network 3
   "Geen Robot Signaal" := "RobotConnectionDB".Stop_value < 1;
   "Noodstop" := "Geen Robot Signaal" OR NOT "Noodstop_aan_Plc" OR NOT "Noodstop_extern";
   IF "Noodstop" THEN
       "HMI_pneumatiek_aan" := FALSE;
       "Tray_Found" := FALSE;
   END_IF;
END_REGION

REGION Network 4
   "Set_Noodstop"();
END_REGION

REGION Network 5
   "RobotConnection"();
END_REGION

REGION Network 6
   "F_TRIG_DB"(CLK := "Noodstop", Q => "HardReset");   // F_TRIG
END_REGION

REGION Network 7
   IF "HardReset" THEN "Reset"(); END_IF;
END_REGION

REGION Network 8
   "Status_Update"();
END_REGION

REGION Network 9
   IF "Running" AND "Pause_Knop" THEN
       "Paused" := TRUE;
       "Tray_Found" := FALSE;
   END_IF;
END_REGION

REGION Network 10
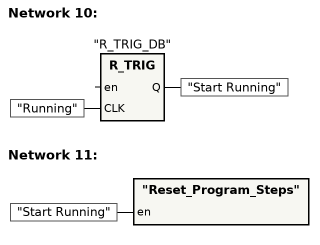
   "R_TRIG_DB"(CLK := "Running", Q => "Start Running");   // R_TRIG
END_REGION

REGION Network 11
   IF "Start Running" THEN "Reset_Program_Steps"(); END_IF;
END_REGION
END_ORGANIZATION_BLOCK

ORGANIZATION_BLOCK "Startup"   // OB100, SCL, Startup
TITLE = "Complete Restart"
{ S7_Optimized_Access := 'FALSE' }
VERSION : 0.1
BEGIN
   //Set Outputs to zero
   "Tafel_uitklappen_cylinder" := 0;
   "Tafel_omhoog_cylinder" := 0;
   "Pneumatiek_aan" := 0;
   "Doosklem_Voor" := 0;
   "Doosklem_Achter" := 0;
   "VAN_ONDEREEEEEN!!!" := 0;

   //Prepare Memory
   "Running" := 0;
   "Noodrestart" := 0;
   "Tafel_hoog" := 0;
   "Next_Box_Ready" := 0;
   "Tray_Found" := 0;
   "Skip Camera" := 0;

   //Prepare Program Steps
   "Waiting for Box" := 1;
   "Box Arrived" := 0;
   "Box Clamped" := 0;
   "Preparing Table" := 0;
   "Waiting for Robot" := 0;
   "Robot is Finished" := 0;
   "!LET HER RIP!" := 0;
END_ORGANIZATION_BLOCK